recipe "Rezeptur": tool_name <- "DB_MouldEditor_HMI_uData_uTools_tool_name", PartShot_Amount <- "DB_MouldEditor_HMI_uData_uTools_PartShot_Amount", RefComponent <- "DB_MouldEditor_HMI_uData_uTools_RefComponent", Spare <- "DB_MouldEditor_HMI_uData_uTools_Spare", EnableTool <- "DB_MouldEditor_HMI_uData_uTools_EnableTool", Spare5_2 <- "DB_MouldEditor_HMI_uData_uTools_Spare5_2", Spare5_3 <- "DB_MouldEditor_HMI_uData_uTools_Spare5_3", Spare5_4 <- "DB_MouldEditor_HMI_uData_uTools_Spare5_4", Spare5_5 <- "DB_MouldEditor_HMI_uData_uTools_Spare5_5", Spare5_6 <- "DB_MouldEditor_HMI_uData_uTools_Spare5_6", EnablePurgeMH <- "DB_MouldEditor_HMI_uData_uTools_EnablePurgeMH", NitrogenVol <- "DB_MouldEditor_HMI_uData_uTools_NitrogenVol", Spare_12 <- "DB_MouldEditor_HMI_uData_uTools_Spare_12", Rob_Prog <- "DB_MouldEditor_HMI_uData_uTools_Rob_Prog", Rob_Prog2 <- "DB_MouldEditor_HMI_uData_uTools_Rob_Prog2", iShotTime <- "DB_MouldEditor_HMI_uData_sColumn_iShotTime", iTotalFlow <- "DB_MouldEditor_HMI_uData_sColumn_iTotalFlow", iTotalWeight <- "DB_MouldEditor_HMI_uData_sColumn_iTotalWeight", arChangePartialShot[0] <- "DB_MouldEditor_HMI_uData_sRow_arChangePartialShot{0}", arChangePartialShot[1] <- "DB_MouldEditor_HMI_uData_sRow_arChangePartialShot{1}", arChangePartialShot[2] <- "DB_MouldEditor_HMI_uData_sRow_arChangePartialShot{2}", arChangePartialShot[3] <- "DB_MouldEditor_HMI_uData_sRow_arChangePartialShot{3}", arChangePartialShot[4] <- "DB_MouldEditor_HMI_uData_sRow_arChangePartialShot{4}", arChangePartialShot[5] <- "DB_MouldEditor_HMI_uData_sRow_arChangePartialShot{5}", arChangePartialShot[6] <- "DB_MouldEditor_HMI_uData_sRow_arChangePartialShot{6}", arChangePartialShot[7] <- "DB_MouldEditor_HMI_uData_sRow_arChangePartialShot{7}", arChangePartialShot[8] <- "DB_MouldEditor_HMI_uData_sRow_arChangePartialShot{8}", arTotalFlow[0] <- "DB_MouldEditor_HMI_uData_sCalculatedValues_arTotalFlow{0}", arTotalFlow[1] <- "DB_MouldEditor_HMI_uData_sCalculatedValues_arTotalFlow{1}", arTotalFlow[2] <- "DB_MouldEditor_HMI_uData_sCalculatedValues_arTotalFlow{2}", arTotalFlow[3] <- "DB_MouldEditor_HMI_uData_sCalculatedValues_arTotalFlow{3}", arTotalFlow[4] <- "DB_MouldEditor_HMI_uData_sCalculatedValues_arTotalFlow{4}", arTotalFlow[5] <- "DB_MouldEditor_HMI_uData_sCalculatedValues_arTotalFlow{5}", arTotalFlow[6] <- "DB_MouldEditor_HMI_uData_sCalculatedValues_arTotalFlow{6}", arTotalFlow[7] <- "DB_MouldEditor_HMI_uData_sCalculatedValues_arTotalFlow{7}", arTotalFlow[8] <- "DB_MouldEditor_HMI_uData_sCalculatedValues_arTotalFlow{8}", MHNo <- "DB_MouldEditor_HMI_uData_arShotSet{0}_MHNo", FoamingTime <- "DB_MouldEditor_HMI_uData_arShotSet{0}_FoamingTime", PartWeight <- "DB_MouldEditor_HMI_uData_arShotSet{0}_PartWeight", CP_ThrottleGap <- "DB_MouldEditor_HMI_uData_arShotSet{0}_CP_ThrottleGap", SwitchOff_Pressure <- "DB_MouldEditor_HMI_uData_arShotSet{0}_SwitchOff_Pressure", PartCounter <- "DB_MouldEditor_HMI_uData_arShotSet{0}_PartCounter", DB_MouldEditor_HMI_uData_arShotSet{0}_RefComponent <- "DB_MouldEditor_HMI_uData_arShotSet{0}_RefComponent", DB_MouldEditor_HMI_uData_arShotSet{0}_PartShotDisable <- "DB_MouldEditor_HMI_uData_arShotSet{0}_PartShotDisable", DB_MouldEditor_HMI_uData_arShotSet{0}_CPMoveAfterShot <- "DB_MouldEditor_HMI_uData_arShotSet{0}_CPMoveAfterShot", DB_MouldEditor_HMI_uData_arShotSet{0}_PurgeMHAfterShot <- "DB_MouldEditor_HMI_uData_arShotSet{0}_PurgeMHAfterShot", DB_MouldEditor_HMI_uData_arShotSet{0}_2PoinMovement_Comp01 <- "DB_MouldEditor_HMI_uData_arShotSet{0}_2PoinMovement_Comp01", DB_MouldEditor_HMI_uData_arShotSet{0}_2PoinMovement_Comp02 <- "DB_MouldEditor_HMI_uData_arShotSet{0}_2PoinMovement_Comp02", DB_MouldEditor_HMI_uData_arShotSet{0}_2PoinMovement_Comp03 <- "DB_MouldEditor_HMI_uData_arShotSet{0}_2PoinMovement_Comp03", DB_MouldEditor_HMI_uData_arShotSet{0}_2PoinMovement_Comp04 <- "DB_MouldEditor_HMI_uData_arShotSet{0}_2PoinMovement_Comp04", DB_MouldEditor_HMI_uData_arShotSet{0}_2PoinMovement_Comp05 <- "DB_MouldEditor_HMI_uData_arShotSet{0}_2PoinMovement_Comp05", DB_MouldEditor_HMI_uData_arShotSet{0}_2PoinMovement_Comp06 <- "DB_MouldEditor_HMI_uData_arShotSet{0}_2PoinMovement_Comp06", DB_MouldEditor_HMI_uData_arShotSet{0}_Spare_1 <- "DB_MouldEditor_HMI_uData_arShotSet{0}_Spare_1", DB_MouldEditor_HMI_uData_arShotSet{0}_Spare_2 <- "DB_MouldEditor_HMI_uData_arShotSet{0}_Spare_2", DB_MouldEditor_HMI_uData_arShotSet{0}_Spare_3 <- "DB_MouldEditor_HMI_uData_arShotSet{0}_Spare_3", DB_MouldEditor_HMI_uData_arShotSet{0}_Spare_4 <- "DB_MouldEditor_HMI_uData_arShotSet{0}_Spare_4", DB_MouldEditor_HMI_uData_arShotSet{0}_Spare_5 <- "DB_MouldEditor_HMI_uData_arShotSet{0}_Spare_5", DB_MouldEditor_HMI_uData_arShotSet{0}_Spare_6 <- "DB_MouldEditor_HMI_uData_arShotSet{0}_Spare_6", DB_MouldEditor_HMI_uData_arShotSet{0}_Spare_7 <- "DB_MouldEditor_HMI_uData_arShotSet{0}_Spare_7", DB_MouldEditor_HMI.uData.arShotSet[1].MHNo <- "DB_MouldEditor_HMI_uData_arShotSet{1}_MHNo", DB_MouldEditor_HMI.uData.arShotSet[1].FoamingTime <- "DB_MouldEditor_HMI_uData_arShotSet{1}_FoamingTime", DB_MouldEditor_HMI.uData.arShotSet[1].PartWeight <- "DB_MouldEditor_HMI_uData_arShotSet{1}_PartWeight", DB_MouldEditor_HMI_uData_arShotSet{1}_CP_ThrottleGap <- "DB_MouldEditor_HMI_uData_arShotSet{1}_CP_ThrottleGap", DB_MouldEditor_HMI_uData_arShotSet{1}_SwitchOff_Pressure <- "DB_MouldEditor_HMI_uData_arShotSet{1}_SwitchOff_Pressure", DB_MouldEditor_HMI.uData.arShotSet[1].PartCounter <- "DB_MouldEditor_HMI_uData_arShotSet{1}_PartCounter", DB_MouldEditor_HMI_uData_arShotSet{1}_RefComponent <- "DB_MouldEditor_HMI_uData_arShotSet{1}_RefComponent", DB_MouldEditor_HMI.uData.arShotSet[1].PartShotDisable <- "DB_MouldEditor_HMI_uData_arShotSet{1}_PartShotDisable", DB_MouldEditor_HMI.uData.arShotSet[1].PurgeMHAfterShot <- "DB_MouldEditor_HMI_uData_arShotSet{1}_PurgeMHAfterShot", DB_MouldEditor_HMI_uData_arShotSet{1}_2PoinMovement_Comp01 <- "DB_MouldEditor_HMI_uData_arShotSet{1}_2PoinMovement_Comp01", DB_MouldEditor_HMI_uData_arShotSet{1}_2PoinMovement_Comp02 <- "DB_MouldEditor_HMI_uData_arShotSet{1}_2PoinMovement_Comp02", DB_MouldEditor_HMI_uData_arShotSet{1}_2PoinMovement_Comp03 <- "DB_MouldEditor_HMI_uData_arShotSet{1}_2PoinMovement_Comp03", DB_MouldEditor_HMI_uData_arShotSet{1}_2PoinMovement_Comp04 <- "DB_MouldEditor_HMI_uData_arShotSet{1}_2PoinMovement_Comp04", DB_MouldEditor_HMI_uData_arShotSet{1}_2PoinMovement_Comp05 <- "DB_MouldEditor_HMI_uData_arShotSet{1}_2PoinMovement_Comp05", DB_MouldEditor_HMI_uData_arShotSet{1}_2PoinMovement_Comp06 <- "DB_MouldEditor_HMI_uData_arShotSet{1}_2PoinMovement_Comp06", DB_MouldEditor_HMI_uData_arShotSet{1}_Spare_1 <- "DB_MouldEditor_HMI_uData_arShotSet{1}_Spare_1", DB_MouldEditor_HMI_uData_arShotSet{1}_Spare_2 <- "DB_MouldEditor_HMI_uData_arShotSet{1}_Spare_2", DB_MouldEditor_HMI_uData_arShotSet{1}_Spare_3 <- "DB_MouldEditor_HMI_uData_arShotSet{1}_Spare_3", DB_MouldEditor_HMI_uData_arShotSet{1}_Spare_4 <- "DB_MouldEditor_HMI_uData_arShotSet{1}_Spare_4", DB_MouldEditor_HMI_uData_arShotSet{1}_Spare_5 <- "DB_MouldEditor_HMI_uData_arShotSet{1}_Spare_5", DB_MouldEditor_HMI_uData_arShotSet{1}_Spare_6 <- "DB_MouldEditor_HMI_uData_arShotSet{1}_Spare_6", DB_MouldEditor_HMI_uData_arShotSet{1}_Spare_7 <- "DB_MouldEditor_HMI_uData_arShotSet{1}_Spare_7", DB_MouldEditor_HMI.uData.arShotSet[2].MHNo <- "DB_MouldEditor_HMI_uData_arShotSet{2}_MHNo", DB_MouldEditor_HMI.uData.arShotSet[2].FoamingTime <- "DB_MouldEditor_HMI_uData_arShotSet{2}_FoamingTime", DB_MouldEditor_HMI.uData.arShotSet[2].PartWeight <- "DB_MouldEditor_HMI_uData_arShotSet{2}_PartWeight", DB_MouldEditor_HMI_uData_arShotSet{2}_CP_ThrottleGap <- "DB_MouldEditor_HMI_uData_arShotSet{2}_CP_ThrottleGap", DB_MouldEditor_HMI_uData_arShotSet{2}_SwitchOff_Pressure <- "DB_MouldEditor_HMI_uData_arShotSet{2}_SwitchOff_Pressure", DB_MouldEditor_HMI.uData.arShotSet[2].PartCounter <- "DB_MouldEditor_HMI_uData_arShotSet{2}_PartCounter", DB_MouldEditor_HMI_uData_arShotSet{2}_RefComponent <- "DB_MouldEditor_HMI_uData_arShotSet{2}_RefComponent", DB_MouldEditor_HMI.uData.arShotSet[2].PartShotDisable <- "DB_MouldEditor_HMI_uData_arShotSet{2}_PartShotDisable", DB_MouldEditor_HMI.uData.arShotSet[2].CPMoveAfterShot <- "DB_MouldEditor_HMI_uData_arShotSet{2}_CPMoveAfterShot", DB_MouldEditor_HMI.uData.arShotSet[2].PurgeMHAfterShot <- "DB_MouldEditor_HMI_uData_arShotSet{2}_PurgeMHAfterShot", DB_MouldEditor_HMI_uData_arShotSet{2}_2PoinMovement_Comp01 <- "DB_MouldEditor_HMI_uData_arShotSet{2}_2PoinMovement_Comp01", DB_MouldEditor_HMI_uData_arShotSet{2}_2PoinMovement_Comp02 <- "DB_MouldEditor_HMI_uData_arShotSet{2}_2PoinMovement_Comp02", DB_MouldEditor_HMI_uData_arShotSet{2}_2PoinMovement_Comp03 <- "DB_MouldEditor_HMI_uData_arShotSet{2}_2PoinMovement_Comp03", DB_MouldEditor_HMI_uData_arShotSet{2}_2PoinMovement_Comp04 <- "DB_MouldEditor_HMI_uData_arShotSet{2}_2PoinMovement_Comp04", DB_MouldEditor_HMI_uData_arShotSet{2}_2PoinMovement_Comp05 <- "DB_MouldEditor_HMI_uData_arShotSet{2}_2PoinMovement_Comp05", DB_MouldEditor_HMI_uData_arShotSet{2}_2PoinMovement_Comp06 <- "DB_MouldEditor_HMI_uData_arShotSet{2}_2PoinMovement_Comp06", DB_MouldEditor_HMI_uData_arShotSet{2}_Spare_1 <- "DB_MouldEditor_HMI_uData_arShotSet{2}_Spare_1", DB_MouldEditor_HMI_uData_arShotSet{2}_Spare_2 <- "DB_MouldEditor_HMI_uData_arShotSet{2}_Spare_2", DB_MouldEditor_HMI_uData_arShotSet{2}_Spare_3 <- "DB_MouldEditor_HMI_uData_arShotSet{2}_Spare_3", DB_MouldEditor_HMI_uData_arShotSet{2}_Spare_4 <- "DB_MouldEditor_HMI_uData_arShotSet{2}_Spare_4", DB_MouldEditor_HMI_uData_arShotSet{2}_Spare_5 <- "DB_MouldEditor_HMI_uData_arShotSet{2}_Spare_5", DB_MouldEditor_HMI_uData_arShotSet{2}_Spare_6 <- "DB_MouldEditor_HMI_uData_arShotSet{2}_Spare_6", DB_MouldEditor_HMI_uData_arShotSet{2}_Spare_7 <- "DB_MouldEditor_HMI_uData_arShotSet{2}_Spare_7", DB_MouldEditor_HMI.uData.arShotSet[3].MHNo <- "DB_MouldEditor_HMI_uData_arShotSet{3}_MHNo", DB_MouldEditor_HMI.uData.arShotSet[3].FoamingTime <- "DB_MouldEditor_HMI_uData_arShotSet{3}_FoamingTime", DB_MouldEditor_HMI.uData.arShotSet[3].PartWeight <- "DB_MouldEditor_HMI_uData_arShotSet{3}_PartWeight", DB_MouldEditor_HMI_uData_arShotSet{3}_CP_ThrottleGap <- "DB_MouldEditor_HMI_uData_arShotSet{3}_CP_ThrottleGap", DB_MouldEditor_HMI_uData_arShotSet{3}_SwitchOff_Pressure <- "DB_MouldEditor_HMI_uData_arShotSet{3}_SwitchOff_Pressure", DB_MouldEditor_HMI.uData.arShotSet[3].PartCounter <- "DB_MouldEditor_HMI_uData_arShotSet{3}_PartCounter", DB_MouldEditor_HMI_uData_arShotSet{3}_RefComponent <- "DB_MouldEditor_HMI_uData_arShotSet{3}_RefComponent", DB_MouldEditor_HMI.uData.arShotSet[3].PartShotDisable <- "DB_MouldEditor_HMI_uData_arShotSet{3}_PartShotDisable", DB_MouldEditor_HMI.uData.arShotSet[3].CPMoveAfterShot <- "DB_MouldEditor_HMI_uData_arShotSet{3}_CPMoveAfterShot", DB_MouldEditor_HMI.uData.arShotSet[3].PurgeMHAfterShot <- "DB_MouldEditor_HMI_uData_arShotSet{3}_PurgeMHAfterShot", DB_MouldEditor_HMI_uData_arShotSet{3}_2PoinMovement_Comp01 <- "DB_MouldEditor_HMI_uData_arShotSet{3}_2PoinMovement_Comp01", DB_MouldEditor_HMI_uData_arShotSet{3}_2PoinMovement_Comp02 <- "DB_MouldEditor_HMI_uData_arShotSet{3}_2PoinMovement_Comp02", DB_MouldEditor_HMI_uData_arShotSet{3}_2PoinMovement_Comp03 <- "DB_MouldEditor_HMI_uData_arShotSet{3}_2PoinMovement_Comp03", DB_MouldEditor_HMI_uData_arShotSet{3}_2PoinMovement_Comp04 <- "DB_MouldEditor_HMI_uData_arShotSet{3}_2PoinMovement_Comp04", DB_MouldEditor_HMI_uData_arShotSet{3}_2PoinMovement_Comp05 <- "DB_MouldEditor_HMI_uData_arShotSet{3}_2PoinMovement_Comp05", DB_MouldEditor_HMI_uData_arShotSet{3}_2PoinMovement_Comp06 <- "DB_MouldEditor_HMI_uData_arShotSet{3}_2PoinMovement_Comp06", DB_MouldEditor_HMI_uData_arShotSet{3}_Spare_1 <- "DB_MouldEditor_HMI_uData_arShotSet{3}_Spare_1", DB_MouldEditor_HMI_uData_arShotSet{3}_Spare_2 <- "DB_MouldEditor_HMI_uData_arShotSet{3}_Spare_2", DB_MouldEditor_HMI_uData_arShotSet{3}_Spare_3 <- "DB_MouldEditor_HMI_uData_arShotSet{3}_Spare_3", DB_MouldEditor_HMI_uData_arShotSet{3}_Spare_4 <- "DB_MouldEditor_HMI_uData_arShotSet{3}_Spare_4", DB_MouldEditor_HMI_uData_arShotSet{3}_Spare_5 <- "DB_MouldEditor_HMI_uData_arShotSet{3}_Spare_5", DB_MouldEditor_HMI_uData_arShotSet{3}_Spare_6 <- "DB_MouldEditor_HMI_uData_arShotSet{3}_Spare_6", DB_MouldEditor_HMI_uData_arShotSet{3}_Spare_7 <- "DB_MouldEditor_HMI_uData_arShotSet{3}_Spare_7", DB_MouldEditor_HMI.uData.arShotSet[4].MHNo <- "DB_MouldEditor_HMI_uData_arShotSet{4}_MHNo", DB_MouldEditor_HMI.uData.arShotSet[4].FoamingTime <- "DB_MouldEditor_HMI_uData_arShotSet{4}_FoamingTime", DB_MouldEditor_HMI.uData.arShotSet[4].PartWeight <- "DB_MouldEditor_HMI_uData_arShotSet{4}_PartWeight", DB_MouldEditor_HMI_uData_arShotSet{4}_CP_ThrottleGap <- "DB_MouldEditor_HMI_uData_arShotSet{4}_CP_ThrottleGap", DB_MouldEditor_HMI_uData_arShotSet{4}_SwitchOff_Pressure <- "DB_MouldEditor_HMI_uData_arShotSet{4}_SwitchOff_Pressure", DB_MouldEditor_HMI.uData.arShotSet[4].PartCounter <- "DB_MouldEditor_HMI_uData_arShotSet{4}_PartCounter", DB_MouldEditor_HMI_uData_arShotSet{4}_RefComponent <- "DB_MouldEditor_HMI_uData_arShotSet{4}_RefComponent", DB_MouldEditor_HMI.uData.arShotSet[4].PartShotDisable <- "DB_MouldEditor_HMI_uData_arShotSet{4}_PartShotDisable", DB_MouldEditor_HMI.uData.arShotSet[4].CPMoveAfterShot <- "DB_MouldEditor_HMI_uData_arShotSet{4}_CPMoveAfterShot", DB_MouldEditor_HMI.uData.arShotSet[4].PurgeMHAfterShot <- "DB_MouldEditor_HMI_uData_arShotSet{4}_PurgeMHAfterShot", DB_MouldEditor_HMI_uData_arShotSet{4}_2PoinMovement_Comp01 <- "DB_MouldEditor_HMI_uData_arShotSet{4}_2PoinMovement_Comp01", DB_MouldEditor_HMI_uData_arShotSet{4}_2PoinMovement_Comp02 <- "DB_MouldEditor_HMI_uData_arShotSet{4}_2PoinMovement_Comp02", DB_MouldEditor_HMI_uData_arShotSet{4}_2PoinMovement_Comp03 <- "DB_MouldEditor_HMI_uData_arShotSet{4}_2PoinMovement_Comp03", DB_MouldEditor_HMI_uData_arShotSet{4}_2PoinMovement_Comp04 <- "DB_MouldEditor_HMI_uData_arShotSet{4}_2PoinMovement_Comp04", DB_MouldEditor_HMI_uData_arShotSet{4}_2PoinMovement_Comp05 <- "DB_MouldEditor_HMI_uData_arShotSet{4}_2PoinMovement_Comp05", DB_MouldEditor_HMI_uData_arShotSet{4}_2PoinMovement_Comp06 <- "DB_MouldEditor_HMI_uData_arShotSet{4}_2PoinMovement_Comp06", DB_MouldEditor_HMI_uData_arShotSet{4}_Spare_1 <- "DB_MouldEditor_HMI_uData_arShotSet{4}_Spare_1", DB_MouldEditor_HMI_uData_arShotSet{4}_Spare_2 <- "DB_MouldEditor_HMI_uData_arShotSet{4}_Spare_2", DB_MouldEditor_HMI_uData_arShotSet{4}_Spare_3 <- "DB_MouldEditor_HMI_uData_arShotSet{4}_Spare_3", DB_MouldEditor_HMI_uData_arShotSet{4}_Spare_4 <- "DB_MouldEditor_HMI_uData_arShotSet{4}_Spare_4", DB_MouldEditor_HMI_uData_arShotSet{4}_Spare_5 <- "DB_MouldEditor_HMI_uData_arShotSet{4}_Spare_5", DB_MouldEditor_HMI_uData_arShotSet{4}_Spare_6 <- "DB_MouldEditor_HMI_uData_arShotSet{4}_Spare_6", DB_MouldEditor_HMI_uData_arShotSet{4}_Spare_7 <- "DB_MouldEditor_HMI_uData_arShotSet{4}_Spare_7", DB_MouldEditor_HMI.uData.arShotSet[5].MHNo <- "DB_MouldEditor_HMI_uData_arShotSet{5}_MHNo", DB_MouldEditor_HMI.uData.arShotSet[5].FoamingTime <- "DB_MouldEditor_HMI_uData_arShotSet{5}_FoamingTime", DB_MouldEditor_HMI.uData.arShotSet[5].PartWeight <- "DB_MouldEditor_HMI_uData_arShotSet{5}_PartWeight", DB_MouldEditor_HMI_uData_arShotSet{5}_CP_ThrottleGap <- "DB_MouldEditor_HMI_uData_arShotSet{5}_CP_ThrottleGap", DB_MouldEditor_HMI_uData_arShotSet{5}_SwitchOff_Pressure <- "DB_MouldEditor_HMI_uData_arShotSet{5}_SwitchOff_Pressure", DB_MouldEditor_HMI.uData.arShotSet[5].PartCounter <- "DB_MouldEditor_HMI_uData_arShotSet{5}_PartCounter", DB_MouldEditor_HMI_uData_arShotSet{5}_RefComponent <- "DB_MouldEditor_HMI_uData_arShotSet{5}_RefComponent", DB_MouldEditor_HMI.uData.arShotSet[5].PartShotDisable <- "DB_MouldEditor_HMI_uData_arShotSet{5}_PartShotDisable", DB_MouldEditor_HMI.uData.arShotSet[5].CPMoveAfterShot <- "DB_MouldEditor_HMI_uData_arShotSet{5}_CPMoveAfterShot", DB_MouldEditor_HMI.uData.arShotSet[5].PurgeMHAfterShot <- "DB_MouldEditor_HMI_uData_arShotSet{5}_PurgeMHAfterShot", DB_MouldEditor_HMI_uData_arShotSet{5}_2PoinMovement_Comp01 <- "DB_MouldEditor_HMI_uData_arShotSet{5}_2PoinMovement_Comp01", DB_MouldEditor_HMI_uData_arShotSet{5}_2PoinMovement_Comp02 <- "DB_MouldEditor_HMI_uData_arShotSet{5}_2PoinMovement_Comp02", DB_MouldEditor_HMI_uData_arShotSet{5}_2PoinMovement_Comp03 <- "DB_MouldEditor_HMI_uData_arShotSet{5}_2PoinMovement_Comp03", DB_MouldEditor_HMI_uData_arShotSet{5}_2PoinMovement_Comp04 <- "DB_MouldEditor_HMI_uData_arShotSet{5}_2PoinMovement_Comp04", DB_MouldEditor_HMI_uData_arShotSet{5}_2PoinMovement_Comp05 <- "DB_MouldEditor_HMI_uData_arShotSet{5}_2PoinMovement_Comp05", DB_MouldEditor_HMI_uData_arShotSet{5}_2PoinMovement_Comp06 <- "DB_MouldEditor_HMI_uData_arShotSet{5}_2PoinMovement_Comp06", DB_MouldEditor_HMI_uData_arShotSet{5}_Spare_1 <- "DB_MouldEditor_HMI_uData_arShotSet{5}_Spare_1", DB_MouldEditor_HMI_uData_arShotSet{5}_Spare_2 <- "DB_MouldEditor_HMI_uData_arShotSet{5}_Spare_2", DB_MouldEditor_HMI_uData_arShotSet{5}_Spare_3 <- "DB_MouldEditor_HMI_uData_arShotSet{5}_Spare_3", DB_MouldEditor_HMI_uData_arShotSet{5}_Spare_4 <- "DB_MouldEditor_HMI_uData_arShotSet{5}_Spare_4", DB_MouldEditor_HMI_uData_arShotSet{5}_Spare_5 <- "DB_MouldEditor_HMI_uData_arShotSet{5}_Spare_5", DB_MouldEditor_HMI_uData_arShotSet{5}_Spare_6 <- "DB_MouldEditor_HMI_uData_arShotSet{5}_Spare_6", DB_MouldEditor_HMI_uData_arShotSet{5}_Spare_7 <- "DB_MouldEditor_HMI_uData_arShotSet{5}_Spare_7", DB_MouldEditor_HMI.uData.arShotSet[6].MHNo <- "DB_MouldEditor_HMI_uData_arShotSet{6}_MHNo", DB_MouldEditor_HMI.uData.arShotSet[6].FoamingTime <- "DB_MouldEditor_HMI_uData_arShotSet{6}_FoamingTime", DB_MouldEditor_HMI.uData.arShotSet[6].PartWeight <- "DB_MouldEditor_HMI_uData_arShotSet{6}_PartWeight", DB_MouldEditor_HMI_uData_arShotSet{6}_CP_ThrottleGap <- "DB_MouldEditor_HMI_uData_arShotSet{6}_CP_ThrottleGap", DB_MouldEditor_HMI_uData_arShotSet{6}_SwitchOff_Pressure <- "DB_MouldEditor_HMI_uData_arShotSet{6}_SwitchOff_Pressure", DB_MouldEditor_HMI.uData.arShotSet[6].PartCounter <- "DB_MouldEditor_HMI_uData_arShotSet{6}_PartCounter", DB_MouldEditor_HMI_uData_arShotSet{6}_RefComponent <- "DB_MouldEditor_HMI_uData_arShotSet{6}_RefComponent", DB_MouldEditor_HMI.uData.arShotSet[6].PartShotDisable <- "DB_MouldEditor_HMI_uData_arShotSet{6}_PartShotDisable", DB_MouldEditor_HMI.uData.arShotSet[6].CPMoveAfterShot <- "DB_MouldEditor_HMI_uData_arShotSet{6}_CPMoveAfterShot", DB_MouldEditor_HMI.uData.arShotSet[6].PurgeMHAfterShot <- "DB_MouldEditor_HMI_uData_arShotSet{6}_PurgeMHAfterShot", DB_MouldEditor_HMI_uData_arShotSet{6}_2PoinMovement_Comp01 <- "DB_MouldEditor_HMI_uData_arShotSet{6}_2PoinMovement_Comp01", DB_MouldEditor_HMI_uData_arShotSet{6}_2PoinMovement_Comp02 <- "DB_MouldEditor_HMI_uData_arShotSet{6}_2PoinMovement_Comp02", DB_MouldEditor_HMI_uData_arShotSet{6}_2PoinMovement_Comp03 <- "DB_MouldEditor_HMI_uData_arShotSet{6}_2PoinMovement_Comp03", DB_MouldEditor_HMI_uData_arShotSet{6}_2PoinMovement_Comp04 <- "DB_MouldEditor_HMI_uData_arShotSet{6}_2PoinMovement_Comp04", DB_MouldEditor_HMI_uData_arShotSet{6}_2PoinMovement_Comp05 <- "DB_MouldEditor_HMI_uData_arShotSet{6}_2PoinMovement_Comp05", DB_MouldEditor_HMI_uData_arShotSet{6}_2PoinMovement_Comp06 <- "DB_MouldEditor_HMI_uData_arShotSet{6}_2PoinMovement_Comp06", DB_MouldEditor_HMI_uData_arShotSet{6}_Spare_1 <- "DB_MouldEditor_HMI_uData_arShotSet{6}_Spare_1", DB_MouldEditor_HMI_uData_arShotSet{6}_Spare_2 <- "DB_MouldEditor_HMI_uData_arShotSet{6}_Spare_2", DB_MouldEditor_HMI_uData_arShotSet{6}_Spare_3 <- "DB_MouldEditor_HMI_uData_arShotSet{6}_Spare_3", DB_MouldEditor_HMI_uData_arShotSet{6}_Spare_4 <- "DB_MouldEditor_HMI_uData_arShotSet{6}_Spare_4", DB_MouldEditor_HMI_uData_arShotSet{6}_Spare_5 <- "DB_MouldEditor_HMI_uData_arShotSet{6}_Spare_5", DB_MouldEditor_HMI_uData_arShotSet{6}_Spare_6 <- "DB_MouldEditor_HMI_uData_arShotSet{6}_Spare_6", DB_MouldEditor_HMI_uData_arShotSet{6}_Spare_7 <- "DB_MouldEditor_HMI_uData_arShotSet{6}_Spare_7", DB_MouldEditor_HMI.uData.arShotSet[7].MHNo <- "DB_MouldEditor_HMI_uData_arShotSet{7}_MHNo", DB_MouldEditor_HMI.uData.arShotSet[7].FoamingTime <- "DB_MouldEditor_HMI_uData_arShotSet{7}_FoamingTime", DB_MouldEditor_HMI.uData.arShotSet[7].PartWeight <- "DB_MouldEditor_HMI_uData_arShotSet{7}_PartWeight", DB_MouldEditor_HMI_uData_arShotSet{7}_CP_ThrottleGap <- "DB_MouldEditor_HMI_uData_arShotSet{7}_CP_ThrottleGap", DB_MouldEditor_HMI_uData_arShotSet{7}_SwitchOff_Pressure <- "DB_MouldEditor_HMI_uData_arShotSet{7}_SwitchOff_Pressure", DB_MouldEditor_HMI.uData.arShotSet[7].PartCounter <- "DB_MouldEditor_HMI_uData_arShotSet{7}_PartCounter", DB_MouldEditor_HMI_uData_arShotSet{7}_RefComponent <- "DB_MouldEditor_HMI_uData_arShotSet{7}_RefComponent", DB_MouldEditor_HMI.uData.arShotSet[7].PartShotDisable <- "DB_MouldEditor_HMI_uData_arShotSet{7}_PartShotDisable", DB_MouldEditor_HMI.uData.arShotSet[7].CPMoveAfterShot <- "DB_MouldEditor_HMI_uData_arShotSet{7}_CPMoveAfterShot", DB_MouldEditor_HMI.uData.arShotSet[7].PurgeMHAfterShot <- "DB_MouldEditor_HMI_uData_arShotSet{7}_PurgeMHAfterShot", DB_MouldEditor_HMI_uData_arShotSet{7}_2PoinMovement_Comp01 <- "DB_MouldEditor_HMI_uData_arShotSet{7}_2PoinMovement_Comp01", DB_MouldEditor_HMI_uData_arShotSet{7}_2PoinMovement_Comp02 <- "DB_MouldEditor_HMI_uData_arShotSet{7}_2PoinMovement_Comp02", DB_MouldEditor_HMI_uData_arShotSet{7}_2PoinMovement_Comp03 <- "DB_MouldEditor_HMI_uData_arShotSet{7}_2PoinMovement_Comp03", DB_MouldEditor_HMI_uData_arShotSet{7}_2PoinMovement_Comp04 <- "DB_MouldEditor_HMI_uData_arShotSet{7}_2PoinMovement_Comp04", DB_MouldEditor_HMI_uData_arShotSet{7}_2PoinMovement_Comp05 <- "DB_MouldEditor_HMI_uData_arShotSet{7}_2PoinMovement_Comp05", DB_MouldEditor_HMI_uData_arShotSet{7}_2PoinMovement_Comp06 <- "DB_MouldEditor_HMI_uData_arShotSet{7}_2PoinMovement_Comp06", DB_MouldEditor_HMI_uData_arShotSet{7}_Spare_1 <- "DB_MouldEditor_HMI_uData_arShotSet{7}_Spare_1", DB_MouldEditor_HMI_uData_arShotSet{7}_Spare_2 <- "DB_MouldEditor_HMI_uData_arShotSet{7}_Spare_2", DB_MouldEditor_HMI_uData_arShotSet{7}_Spare_3 <- "DB_MouldEditor_HMI_uData_arShotSet{7}_Spare_3", DB_MouldEditor_HMI_uData_arShotSet{7}_Spare_4 <- "DB_MouldEditor_HMI_uData_arShotSet{7}_Spare_4", DB_MouldEditor_HMI_uData_arShotSet{7}_Spare_5 <- "DB_MouldEditor_HMI_uData_arShotSet{7}_Spare_5", DB_MouldEditor_HMI_uData_arShotSet{7}_Spare_6 <- "DB_MouldEditor_HMI_uData_arShotSet{7}_Spare_6", DB_MouldEditor_HMI_uData_arShotSet{7}_Spare_7 <- "DB_MouldEditor_HMI_uData_arShotSet{7}_Spare_7", DB_MouldEditor_HMI.uData.arShotSet[8].MHNo <- "DB_MouldEditor_HMI_uData_arShotSet{8}_MHNo", DB_MouldEditor_HMI.uData.arShotSet[8].FoamingTime <- "DB_MouldEditor_HMI_uData_arShotSet{8}_FoamingTime", DB_MouldEditor_HMI.uData.arShotSet[8].PartWeight <- "DB_MouldEditor_HMI_uData_arShotSet{8}_PartWeight", DB_MouldEditor_HMI_uData_arShotSet{8}_CP_ThrottleGap <- "DB_MouldEditor_HMI_uData_arShotSet{8}_CP_ThrottleGap", DB_MouldEditor_HMI_uData_arShotSet{8}_SwitchOff_Pressure <- "DB_MouldEditor_HMI_uData_arShotSet{8}_SwitchOff_Pressure", DB_MouldEditor_HMI.uData.arShotSet[8].PartCounter <- "DB_MouldEditor_HMI_uData_arShotSet{8}_PartCounter", DB_MouldEditor_HMI_uData_arShotSet{8}_RefComponent <- "DB_MouldEditor_HMI_uData_arShotSet{8}_RefComponent", DB_MouldEditor_HMI.uData.arShotSet[8].PartShotDisable <- "DB_MouldEditor_HMI_uData_arShotSet{8}_PartShotDisable", DB_MouldEditor_HMI.uData.arShotSet[8].CPMoveAfterShot <- "DB_MouldEditor_HMI_uData_arShotSet{8}_CPMoveAfterShot", DB_MouldEditor_HMI.uData.arShotSet[8].PurgeMHAfterShot <- "DB_MouldEditor_HMI_uData_arShotSet{8}_PurgeMHAfterShot", DB_MouldEditor_HMI_uData_arShotSet{8}_2PoinMovement_Comp01 <- "DB_MouldEditor_HMI_uData_arShotSet{8}_2PoinMovement_Comp01", DB_MouldEditor_HMI_uData_arShotSet{8}_2PoinMovement_Comp02 <- "DB_MouldEditor_HMI_uData_arShotSet{8}_2PoinMovement_Comp02", DB_MouldEditor_HMI_uData_arShotSet{8}_2PoinMovement_Comp03 <- "DB_MouldEditor_HMI_uData_arShotSet{8}_2PoinMovement_Comp03", DB_MouldEditor_HMI_uData_arShotSet{8}_2PoinMovement_Comp04 <- "DB_MouldEditor_HMI_uData_arShotSet{8}_2PoinMovement_Comp04", DB_MouldEditor_HMI_uData_arShotSet{8}_2PoinMovement_Comp05 <- "DB_MouldEditor_HMI_uData_arShotSet{8}_2PoinMovement_Comp05", DB_MouldEditor_HMI_uData_arShotSet{8}_2PoinMovement_Comp06 <- "DB_MouldEditor_HMI_uData_arShotSet{8}_2PoinMovement_Comp06", DB_MouldEditor_HMI_uData_arShotSet{8}_Spare_1 <- "DB_MouldEditor_HMI_uData_arShotSet{8}_Spare_1", DB_MouldEditor_HMI_uData_arShotSet{8}_Spare_2 <- "DB_MouldEditor_HMI_uData_arShotSet{8}_Spare_2", DB_MouldEditor_HMI_uData_arShotSet{8}_Spare_3 <- "DB_MouldEditor_HMI_uData_arShotSet{8}_Spare_3", DB_MouldEditor_HMI_uData_arShotSet{8}_Spare_4 <- "DB_MouldEditor_HMI_uData_arShotSet{8}_Spare_4", DB_MouldEditor_HMI_uData_arShotSet{8}_Spare_5 <- "DB_MouldEditor_HMI_uData_arShotSet{8}_Spare_5", DB_MouldEditor_HMI_uData_arShotSet{8}_Spare_6 <- "DB_MouldEditor_HMI_uData_arShotSet{8}_Spare_6", DB_MouldEditor_HMI_uData_arShotSet{8}_Spare_7 <- "DB_MouldEditor_HMI_uData_arShotSet{8}_Spare_7", DB_MouldEditor_HMI_uData_arShotSet{0}_Pressure{1} <- "DB_MouldEditor_HMI_uData_arShotSet{0}_Pressure{1}", DB_MouldEditor_HMI_uData_arShotSet{0}_Pressure{2} <- "DB_MouldEditor_HMI_uData_arShotSet{0}_Pressure{2}", DB_MouldEditor_HMI_uData_arShotSet{0}_Pressure{3} <- "DB_MouldEditor_HMI_uData_arShotSet{0}_Pressure{3}", DB_MouldEditor_HMI_uData_arShotSet{0}_Pressure{4} <- "DB_MouldEditor_HMI_uData_arShotSet{0}_Pressure{4}", DB_MouldEditor_HMI_uData_arShotSet{0}_Pressure{5} <- "DB_MouldEditor_HMI_uData_arShotSet{0}_Pressure{5}", DB_MouldEditor_HMI_uData_arShotSet{0}_Pressure{6} <- "DB_MouldEditor_HMI_uData_arShotSet{0}_Pressure{6}", DB_MouldEditor_HMI_uData_arShotSet{0}_Flow{2} <- "DB_MouldEditor_HMI_uData_arShotSet{0}_Flow{2}", DB_MouldEditor_HMI_uData_arShotSet{0}_Flow{1} <- "DB_MouldEditor_HMI_uData_arShotSet{0}_Flow{1}", DB_MouldEditor_HMI_uData_arShotSet{0}_Flow{3} <- "DB_MouldEditor_HMI_uData_arShotSet{0}_Flow{3}", DB_MouldEditor_HMI_uData_arShotSet{0}_Flow{4} <- "DB_MouldEditor_HMI_uData_arShotSet{0}_Flow{4}", DB_MouldEditor_HMI_uData_arShotSet{0}_Flow{5} <- "DB_MouldEditor_HMI_uData_arShotSet{0}_Flow{5}", DB_MouldEditor_HMI_uData_arShotSet{0}_Flow{6} <- "DB_MouldEditor_HMI_uData_arShotSet{0}_Flow{6}", DB_MouldEditor_HMI_uData_arShotSet{1}_Flow{1} <- "DB_MouldEditor_HMI_uData_arShotSet{1}_Flow{1}", DB_MouldEditor_HMI_uData_arShotSet{1}_Flow{2} <- "DB_MouldEditor_HMI_uData_arShotSet{1}_Flow{2}", DB_MouldEditor_HMI_uData_arShotSet{1}_Flow{3} <- "DB_MouldEditor_HMI_uData_arShotSet{1}_Flow{3}", DB_MouldEditor_HMI_uData_arShotSet{1}_Flow{4} <- "DB_MouldEditor_HMI_uData_arShotSet{1}_Flow{4}", DB_MouldEditor_HMI_uData_arShotSet{1}_Flow{5} <- "DB_MouldEditor_HMI_uData_arShotSet{1}_Flow{5}", DB_MouldEditor_HMI_uData_arShotSet{1}_Flow{6} <- "DB_MouldEditor_HMI_uData_arShotSet{1}_Flow{6}", DB_MouldEditor_HMI_uData_arShotSet{1}_Pressure{1} <- "DB_MouldEditor_HMI_uData_arShotSet{1}_Pressure{1}", DB_MouldEditor_HMI_uData_arShotSet{1}_Pressure{2} <- "DB_MouldEditor_HMI_uData_arShotSet{1}_Pressure{2}", DB_MouldEditor_HMI_uData_arShotSet{1}_Pressure{3} <- "DB_MouldEditor_HMI_uData_arShotSet{1}_Pressure{3}", DB_MouldEditor_HMI_uData_arShotSet{1}_Pressure{4} <- "DB_MouldEditor_HMI_uData_arShotSet{1}_Pressure{4}", DB_MouldEditor_HMI_uData_arShotSet{1}_Pressure{5} <- "DB_MouldEditor_HMI_uData_arShotSet{1}_Pressure{5}", DB_MouldEditor_HMI_uData_arShotSet{1}_Pressure{6} <- "DB_MouldEditor_HMI_uData_arShotSet{1}_Pressure{6}", DB_MouldEditor_HMI_uData_arShotSet{2}_Flow{1} <- "DB_MouldEditor_HMI_uData_arShotSet{2}_Flow{1}", DB_MouldEditor_HMI_uData_arShotSet{2}_Flow{2} <- "DB_MouldEditor_HMI_uData_arShotSet{2}_Flow{2}", DB_MouldEditor_HMI_uData_arShotSet{2}_Flow{3} <- "DB_MouldEditor_HMI_uData_arShotSet{2}_Flow{3}", DB_MouldEditor_HMI_uData_arShotSet{2}_Flow{4} <- "DB_MouldEditor_HMI_uData_arShotSet{2}_Flow{4}", DB_MouldEditor_HMI_uData_arShotSet{2}_Flow{5} <- "DB_MouldEditor_HMI_uData_arShotSet{2}_Flow{5}", DB_MouldEditor_HMI_uData_arShotSet{2}_Flow{6} <- "DB_MouldEditor_HMI_uData_arShotSet{2}_Flow{6}", DB_MouldEditor_HMI_uData_arShotSet{2}_Pressure{1} <- "DB_MouldEditor_HMI_uData_arShotSet{2}_Pressure{1}", DB_MouldEditor_HMI_uData_arShotSet{2}_Pressure{2} <- "DB_MouldEditor_HMI_uData_arShotSet{2}_Pressure{2}", DB_MouldEditor_HMI_uData_arShotSet{2}_Pressure{3} <- "DB_MouldEditor_HMI_uData_arShotSet{2}_Pressure{3}", DB_MouldEditor_HMI_uData_arShotSet{2}_Pressure{4} <- "DB_MouldEditor_HMI_uData_arShotSet{2}_Pressure{4}", DB_MouldEditor_HMI_uData_arShotSet{2}_Pressure{5} <- "DB_MouldEditor_HMI_uData_arShotSet{2}_Pressure{5}", DB_MouldEditor_HMI_uData_arShotSet{2}_Pressure{6} <- "DB_MouldEditor_HMI_uData_arShotSet{2}_Pressure{6}", DB_MouldEditor_HMI_uData_arShotSet{3}_Flow{1} <- "DB_MouldEditor_HMI_uData_arShotSet{3}_Flow{1}", DB_MouldEditor_HMI_uData_arShotSet{3}_Flow{2} <- "DB_MouldEditor_HMI_uData_arShotSet{3}_Flow{2}", DB_MouldEditor_HMI_uData_arShotSet{3}_Flow{3} <- "DB_MouldEditor_HMI_uData_arShotSet{3}_Flow{3}", DB_MouldEditor_HMI_uData_arShotSet{3}_Flow{4} <- "DB_MouldEditor_HMI_uData_arShotSet{3}_Flow{4}", DB_MouldEditor_HMI_uData_arShotSet{3}_Flow{5} <- "DB_MouldEditor_HMI_uData_arShotSet{3}_Flow{5}", DB_MouldEditor_HMI_uData_arShotSet{3}_Flow{6} <- "DB_MouldEditor_HMI_uData_arShotSet{3}_Flow{6}", DB_MouldEditor_HMI_uData_arShotSet{3}_Pressure{1} <- "DB_MouldEditor_HMI_uData_arShotSet{3}_Pressure{1}", DB_MouldEditor_HMI_uData_arShotSet{3}_Pressure{2} <- "DB_MouldEditor_HMI_uData_arShotSet{3}_Pressure{2}", DB_MouldEditor_HMI_uData_arShotSet{3}_Pressure{3} <- "DB_MouldEditor_HMI_uData_arShotSet{3}_Pressure{3}", DB_MouldEditor_HMI_uData_arShotSet{3}_Pressure{4} <- "DB_MouldEditor_HMI_uData_arShotSet{3}_Pressure{4}", DB_MouldEditor_HMI_uData_arShotSet{3}_Pressure{5} <- "DB_MouldEditor_HMI_uData_arShotSet{3}_Pressure{5}", DB_MouldEditor_HMI_uData_arShotSet{3}_Pressure{6} <- "DB_MouldEditor_HMI_uData_arShotSet{3}_Pressure{6}", DB_MouldEditor_HMI_uData_arShotSet{4}_Flow{1} <- "DB_MouldEditor_HMI_uData_arShotSet{4}_Flow{1}", DB_MouldEditor_HMI_uData_arShotSet{4}_Flow{2} <- "DB_MouldEditor_HMI_uData_arShotSet{4}_Flow{2}", DB_MouldEditor_HMI_uData_arShotSet{4}_Flow{3} <- "DB_MouldEditor_HMI_uData_arShotSet{4}_Flow{3}", DB_MouldEditor_HMI_uData_arShotSet{4}_Flow{4} <- "DB_MouldEditor_HMI_uData_arShotSet{4}_Flow{4}", DB_MouldEditor_HMI_uData_arShotSet{4}_Flow{5} <- "DB_MouldEditor_HMI_uData_arShotSet{4}_Flow{5}", DB_MouldEditor_HMI_uData_arShotSet{4}_Flow{6} <- "DB_MouldEditor_HMI_uData_arShotSet{4}_Flow{6}", DB_MouldEditor_HMI_uData_arShotSet{4}_Pressure{1} <- "DB_MouldEditor_HMI_uData_arShotSet{4}_Pressure{1}", DB_MouldEditor_HMI_uData_arShotSet{4}_Pressure{2} <- "DB_MouldEditor_HMI_uData_arShotSet{4}_Pressure{2}", DB_MouldEditor_HMI_uData_arShotSet{4}_Pressure{3} <- "DB_MouldEditor_HMI_uData_arShotSet{4}_Pressure{3}", DB_MouldEditor_HMI_uData_arShotSet{4}_Pressure{4} <- "DB_MouldEditor_HMI_uData_arShotSet{4}_Pressure{4}", DB_MouldEditor_HMI_uData_arShotSet{4}_Pressure{5} <- "DB_MouldEditor_HMI_uData_arShotSet{4}_Pressure{5}", DB_MouldEditor_HMI_uData_arShotSet{4}_Pressure{6} <- "DB_MouldEditor_HMI_uData_arShotSet{4}_Pressure{6}", DB_MouldEditor_HMI_uData_arShotSet{5}_Flow{1} <- "DB_MouldEditor_HMI_uData_arShotSet{5}_Flow{1}", DB_MouldEditor_HMI_uData_arShotSet{5}_Flow{2} <- "DB_MouldEditor_HMI_uData_arShotSet{5}_Flow{2}", DB_MouldEditor_HMI_uData_arShotSet{5}_Flow{3} <- "DB_MouldEditor_HMI_uData_arShotSet{5}_Flow{3}", DB_MouldEditor_HMI_uData_arShotSet{5}_Flow{4} <- "DB_MouldEditor_HMI_uData_arShotSet{5}_Flow{4}", DB_MouldEditor_HMI_uData_arShotSet{5}_Flow{5} <- "DB_MouldEditor_HMI_uData_arShotSet{5}_Flow{5}", DB_MouldEditor_HMI_uData_arShotSet{5}_Flow{6} <- "DB_MouldEditor_HMI_uData_arShotSet{5}_Flow{6}", DB_MouldEditor_HMI_uData_arShotSet{5}_Pressure{1} <- "DB_MouldEditor_HMI_uData_arShotSet{5}_Pressure{1}", DB_MouldEditor_HMI_uData_arShotSet{5}_Pressure{2} <- "DB_MouldEditor_HMI_uData_arShotSet{5}_Pressure{2}", DB_MouldEditor_HMI_uData_arShotSet{5}_Pressure{3} <- "DB_MouldEditor_HMI_uData_arShotSet{5}_Pressure{3}", DB_MouldEditor_HMI_uData_arShotSet{5}_Pressure{4} <- "DB_MouldEditor_HMI_uData_arShotSet{5}_Pressure{4}", DB_MouldEditor_HMI_uData_arShotSet{5}_Pressure{5} <- "DB_MouldEditor_HMI_uData_arShotSet{5}_Pressure{5}", DB_MouldEditor_HMI_uData_arShotSet{5}_Pressure{6} <- "DB_MouldEditor_HMI_uData_arShotSet{5}_Pressure{6}", DB_MouldEditor_HMI_uData_arShotSet{6}_Flow{1} <- "DB_MouldEditor_HMI_uData_arShotSet{6}_Flow{1}", DB_MouldEditor_HMI_uData_arShotSet{6}_Flow{2} <- "DB_MouldEditor_HMI_uData_arShotSet{6}_Flow{2}", DB_MouldEditor_HMI_uData_arShotSet{6}_Flow{3} <- "DB_MouldEditor_HMI_uData_arShotSet{6}_Flow{3}", DB_MouldEditor_HMI_uData_arShotSet{6}_Flow{4} <- "DB_MouldEditor_HMI_uData_arShotSet{6}_Flow{4}", DB_MouldEditor_HMI_uData_arShotSet{6}_Flow{5} <- "DB_MouldEditor_HMI_uData_arShotSet{6}_Flow{5}", DB_MouldEditor_HMI_uData_arShotSet{6}_Flow{6} <- "DB_MouldEditor_HMI_uData_arShotSet{6}_Flow{6}", DB_MouldEditor_HMI_uData_arShotSet{6}_Pressure{1} <- "DB_MouldEditor_HMI_uData_arShotSet{6}_Pressure{1}", DB_MouldEditor_HMI_uData_arShotSet{6}_Pressure{2} <- "DB_MouldEditor_HMI_uData_arShotSet{6}_Pressure{2}", DB_MouldEditor_HMI_uData_arShotSet{6}_Pressure{3} <- "DB_MouldEditor_HMI_uData_arShotSet{6}_Pressure{3}", DB_MouldEditor_HMI_uData_arShotSet{6}_Pressure{4} <- "DB_MouldEditor_HMI_uData_arShotSet{6}_Pressure{4}", DB_MouldEditor_HMI_uData_arShotSet{6}_Pressure{5} <- "DB_MouldEditor_HMI_uData_arShotSet{6}_Pressure{5}", DB_MouldEditor_HMI_uData_arShotSet{6}_Pressure{6} <- "DB_MouldEditor_HMI_uData_arShotSet{6}_Pressure{6}", DB_MouldEditor_HMI_uData_arShotSet{7}_Flow{1} <- "DB_MouldEditor_HMI_uData_arShotSet{7}_Flow{1}", DB_MouldEditor_HMI_uData_arShotSet{7}_Flow{2} <- "DB_MouldEditor_HMI_uData_arShotSet{7}_Flow{2}", DB_MouldEditor_HMI_uData_arShotSet{7}_Flow{3} <- "DB_MouldEditor_HMI_uData_arShotSet{7}_Flow{3}", DB_MouldEditor_HMI_uData_arShotSet{7}_Flow{4} <- "DB_MouldEditor_HMI_uData_arShotSet{7}_Flow{4}", DB_MouldEditor_HMI_uData_arShotSet{7}_Flow{5} <- "DB_MouldEditor_HMI_uData_arShotSet{7}_Flow{5}", DB_MouldEditor_HMI_uData_arShotSet{7}_Flow{6} <- "DB_MouldEditor_HMI_uData_arShotSet{7}_Flow{6}", DB_MouldEditor_HMI_uData_arShotSet{7}_Pressure{1} <- "DB_MouldEditor_HMI_uData_arShotSet{7}_Pressure{1}", DB_MouldEditor_HMI_uData_arShotSet{7}_Pressure{2} <- "DB_MouldEditor_HMI_uData_arShotSet{7}_Pressure{2}", DB_MouldEditor_HMI_uData_arShotSet{7}_Pressure{3} <- "DB_MouldEditor_HMI_uData_arShotSet{7}_Pressure{3}", DB_MouldEditor_HMI_uData_arShotSet{7}_Pressure{4} <- "DB_MouldEditor_HMI_uData_arShotSet{7}_Pressure{4}", DB_MouldEditor_HMI_uData_arShotSet{7}_Pressure{5} <- "DB_MouldEditor_HMI_uData_arShotSet{7}_Pressure{5}", DB_MouldEditor_HMI_uData_arShotSet{7}_Pressure{6} <- "DB_MouldEditor_HMI_uData_arShotSet{7}_Pressure{6}", DB_MouldEditor_HMI_uData_arShotSet{8}_Flow{1} <- "DB_MouldEditor_HMI_uData_arShotSet{8}_Flow{1}", DB_MouldEditor_HMI_uData_arShotSet{8}_Flow{2} <- "DB_MouldEditor_HMI_uData_arShotSet{8}_Flow{2}", DB_MouldEditor_HMI_uData_arShotSet{8}_Flow{3} <- "DB_MouldEditor_HMI_uData_arShotSet{8}_Flow{3}", DB_MouldEditor_HMI_uData_arShotSet{8}_Flow{4} <- "DB_MouldEditor_HMI_uData_arShotSet{8}_Flow{4}", DB_MouldEditor_HMI_uData_arShotSet{8}_Flow{5} <- "DB_MouldEditor_HMI_uData_arShotSet{8}_Flow{5}", DB_MouldEditor_HMI_uData_arShotSet{8}_Flow{6} <- "DB_MouldEditor_HMI_uData_arShotSet{8}_Flow{6}", DB_MouldEditor_HMI_uData_arShotSet{8}_Pressure{1} <- "DB_MouldEditor_HMI_uData_arShotSet{8}_Pressure{1}", DB_MouldEditor_HMI_uData_arShotSet{8}_Pressure{2} <- "DB_MouldEditor_HMI_uData_arShotSet{8}_Pressure{2}", DB_MouldEditor_HMI_uData_arShotSet{8}_Pressure{3} <- "DB_MouldEditor_HMI_uData_arShotSet{8}_Pressure{3}", DB_MouldEditor_HMI_uData_arShotSet{8}_Pressure{4} <- "DB_MouldEditor_HMI_uData_arShotSet{8}_Pressure{4}", DB_MouldEditor_HMI_uData_arShotSet{8}_Pressure{5} <- "DB_MouldEditor_HMI_uData_arShotSet{8}_Pressure{5}", DB_MouldEditor_HMI_uData_arShotSet{8}_Pressure{6} <- "DB_MouldEditor_HMI_uData_arShotSet{8}_Pressure{6}", DB_MouldEditor_HMI_uData_sSelected_sPS_arFlow{0} <- "DB_MouldEditor_HMI_uData_sSelected_sPS_arFlow{0}", DB_MouldEditor_HMI_uData_sSelected_sPS_arRatio{0} <- "DB_MouldEditor_HMI_uData_sSelected_sPS_arRatio{0}", DB_MouldEditor_HMI_uData_sSelected_sPS_arPressure{0} <- "DB_MouldEditor_HMI_uData_sSelected_sPS_arPressure{0}", DB_MouldEditor_HMI_uData_sSelected_sPS_2PoinMovement_Comp01 <- "DB_MouldEditor_HMI_uData_sSelected_sPS_2PoinMovement_Comp01", DB_MouldEditor_HMI_uData_sSelected_sPS_2PoinMovement_Comp02 <- "DB_MouldEditor_HMI_uData_sSelected_sPS_2PoinMovement_Comp02", DB_MouldEditor_HMI_uData_sSelected_sPS_2PoinMovement_Comp03 <- "DB_MouldEditor_HMI_uData_sSelected_sPS_2PoinMovement_Comp03", DB_MouldEditor_HMI_uData_sSelected_sPS_2PoinMovement_Comp04 <- "DB_MouldEditor_HMI_uData_sSelected_sPS_2PoinMovement_Comp04", DB_MouldEditor_HMI_uData_sSelected_sPS_2PoinMovement_Comp05 <- "DB_MouldEditor_HMI_uData_sSelected_sPS_2PoinMovement_Comp05", DB_MouldEditor_HMI_uData_sSelected_sPS_2PoinMovement_Comp06 <- "DB_MouldEditor_HMI_uData_sSelected_sPS_2PoinMovement_Comp06", DB_MouldEditor_HMI_uData_sSelected_iCalculation <- "DB_MouldEditor_HMI_uData_sSelected_iCalculation", DB_MouldEditor_HMI_uData_sSelected_iTool <- "DB_MouldEditor_HMI_uData_sSelected_iTool", DB_MouldEditor_HMI_uData_sSelected_sPS_arFlow{1} <- "DB_MouldEditor_HMI_uData_sSelected_sPS_arFlow{1}", DB_MouldEditor_HMI_uData_sSelected_sPS_arFlow{2} <- "DB_MouldEditor_HMI_uData_sSelected_sPS_arFlow{2}", DB_MouldEditor_HMI_uData_sSelected_sPS_arFlow{3} <- "DB_MouldEditor_HMI_uData_sSelected_sPS_arFlow{3}", DB_MouldEditor_HMI_uData_sSelected_sPS_arFlow{4} <- "DB_MouldEditor_HMI_uData_sSelected_sPS_arFlow{4}", DB_MouldEditor_HMI_uData_sSelected_sPS_arFlow{5} <- "DB_MouldEditor_HMI_uData_sSelected_sPS_arFlow{5}", DB_MouldEditor_HMI_uData_sSelected_sPS_arFlow{6} <- "DB_MouldEditor_HMI_uData_sSelected_sPS_arFlow{6}", DB_MouldEditor_HMI_uData_sSelected_sPS_arPressure{1} <- "DB_MouldEditor_HMI_uData_sSelected_sPS_arPressure{1}", DB_MouldEditor_HMI_uData_sSelected_sPS_arPressure{2} <- "DB_MouldEditor_HMI_uData_sSelected_sPS_arPressure{2}", DB_MouldEditor_HMI_uData_sSelected_sPS_arPressure{3} <- "DB_MouldEditor_HMI_uData_sSelected_sPS_arPressure{3}", DB_MouldEditor_HMI_uData_sSelected_sPS_arPressure{4} <- "DB_MouldEditor_HMI_uData_sSelected_sPS_arPressure{4}", DB_MouldEditor_HMI_uData_sSelected_sPS_arPressure{5} <- "DB_MouldEditor_HMI_uData_sSelected_sPS_arPressure{5}", DB_MouldEditor_HMI_uData_sSelected_sPS_arPressure{6} <- "DB_MouldEditor_HMI_uData_sSelected_sPS_arPressure{6}", DB_MouldEditor_HMI_uData_sSelected_sPS_arRatio{1} <- "DB_MouldEditor_HMI_uData_sSelected_sPS_arRatio{1}", DB_MouldEditor_HMI_uData_sSelected_sPS_arRatio{2} <- "DB_MouldEditor_HMI_uData_sSelected_sPS_arRatio{2}", DB_MouldEditor_HMI_uData_sSelected_sPS_arRatio{3} <- "DB_MouldEditor_HMI_uData_sSelected_sPS_arRatio{3}", DB_MouldEditor_HMI_uData_sSelected_sPS_arRatio <- "DB_MouldEditor_HMI_uData_sSelected_sPS_arRatio{4}", DB_MouldEditor_HMI_uData_sSelected_sPS_arRatio{5} <- "DB_MouldEditor_HMI_uData_sSelected_sPS_arRatio{5}", DB_MouldEditor_HMI_uData_sSelected_sPS_arRatio{6} <- "DB_MouldEditor_HMI_uData_sSelected_sPS_arRatio{6}", DB_MouldEditor_HMI_uData_sSelected_sPS_iPS <- "DB_MouldEditor_HMI_uData_sSelected_sPS_iPS", DB_MouldEditor_HMI_uData_sSelected_sPS_RefComponent <- "DB_MouldEditor_HMI_uData_sSelected_sPS_RefComponent"

recipe "Shifttime": Recipe_element_1 <- "Shift_1_1", Recipe_element_2 <- "Shift_1_2", Recipe_element_3 <- "Shift_1_3", Recipe_element_4 <- "Shift_1_4", Recipe_element_5 <- "Shift_2_1", Recipe_element_6 <- "Shift_2_2", Recipe_element_7 <- "Shift_2_3", Recipe_element_8 <- "Shift_2_4", Recipe_element_9 <- "Shift_3_1", Recipe_element_10 <- "Shift_3_2", Recipe_element_11 <- "Shift_3_3", Recipe_element_12 <- "Shift_3_4", Recipe_element_13 <- "Shift_4_1", Recipe_element_14 <- "Shift_4_2", Recipe_element_15 <- "Shift_4_3", Recipe_element_16 <- "Shift_4_4", Recipe_element_17 <- "Shift_5_1", Recipe_element_18 <- "Shift_5_2", Recipe_element_19 <- "Shift_5_3", Recipe_element_20 <- "Shift_5_4", Recipe_element_21 <- "Shift_6_1", Recipe_element_22 <- "Shift_6_2", Recipe_element_23 <- "Shift_6_3", Recipe_element_24 <- "Shift_6_4", Recipe_element_25 <- "Shift_7_1", Recipe_element_26 <- "Shift_7_2", Recipe_element_27 <- "Shift_7_3", Recipe_element_28 <- "Shift_7_4", Recipe_element_29 <- "Shift_En_1_1", Recipe_element_30 <- "Shift_En_1_2", Recipe_element_31 <- "Shift_En_1_3", Recipe_element_32 <- "Shift_En_1_4", Recipe_element_33 <- "Shift_En_2_1", Recipe_element_34 <- "Shift_En_2_2", Recipe_element_35 <- "Shift_En_2_3", Recipe_element_36 <- "Shift_En_2_4", Recipe_element_37 <- "Shift_En_3_1", Recipe_element_38 <- "Shift_En_3_2", Recipe_element_39 <- "Shift_En_3_3", Recipe_element_40 <- "Shift_En_3_4", Recipe_element_41 <- "Shift_En_4_1", Recipe_element_42 <- "Shift_En_4_2", Recipe_element_43 <- "Shift_En_4_3", Recipe_element_44 <- "Shift_En_4_4", Recipe_element_45 <- "Shift_En_5_1", Recipe_element_46 <- "Shift_En_5_2", Recipe_element_47 <- "Shift_En_5_3", Recipe_element_48 <- "Shift_En_5_4", Recipe_element_49 <- "Shift_En_6_1", Recipe_element_50 <- "Shift_En_6_2", Recipe_element_51 <- "Shift_En_6_3", Recipe_element_52 <- "Shift_En_6_4", Recipe_element_53 <- "Shift_En_7_1", Recipe_element_54 <- "Shift_En_7_2", Recipe_element_55 <- "Shift_En_7_3", Recipe_element_56 <- "Shift_En_7_4"

recipe "ShiftProtocol": Shift_Protocol_1 <- "Shift_Protocol_1", Shift_Protocol_2 <- "Shift_Protocol_2", Shift_Protocol_3 <- "Shift_Protocol_3", Shift_Protocol_4 <- "Shift_Protocol_4", Shift_Protocol_5 <- "Shift_Protocol_5", Shift_Protocol_6 <- "Shift_Protocol_6", Shift_Protocol_7 <- "Shift_Protocol_7", Shift_Protocol_8 <- "Shift_Protocol_8", Shift_Protocol_9 <- "Shift_Protocol_9", Shift_Protocol_10 <- "Shift_Protocol_10", Shift_Protocol_11 <- "Shift_Protocol_11", Shift_Protocol_12 <- "Shift_Protocol_12", Shift_Protocol_13 <- "Shift_Protocol_13", Shift_Protocol_14 <- "Shift_Protocol_14", Shift_Protocol_15 <- "Shift_Protocol_15", Shift_Protocol_16 <- "Shift_Protocol_16", Shift_Protocol_17 <- "Shift_Protocol_17", Shift_Protocol_18 <- "Shift_Protocol_18", Shift_Protocol_19 <- "Shift_Protocol_19", Shift_Protocol_20 <- "Shift_Protocol_20", Shift_Protocol_21 <- "Shift_Protocol_21"